(* Logix 5000 project; controller PLC_MCC1300_75F1 vendor 1 type 14 code 166 rev 32.11; software revision 32.04; part 42 of 83 *)
(* tags used below, declared in another part *)
   AUX_xDebugNewPlate : BOOL;
   CM_DATA_Snap_Rx : CM_DATA_Z200;
   CM_INPUT_Z200_Sync : CM_INPUT_Z200;
   CONST_tAux : AUX_COSTANTS;
   CONST_tPlant : UDT_PLANT_CONSTANTS;
   ECL_HLD_AUTO : ALIAS FOR N14[240].2;
   ECL_HLD_AUTO_N : ALIAS FOR I[36].14;
   ECL_HLD_AUTO_S : ALIAS FOR I[80].14;
   ECL_HLD_UP : ALIAS FOR N14[240].3;
   ECL_HLD_UP_N : ALIAS FOR I[36].15;
   ECL_HLD_UP_S : ALIAS FOR I[80].15;
   FL_HLD_AUTO : ALIAS FOR N14[240].0;
   FL_HLD_AUTO_N : ALIAS FOR I[36].12;
   FL_HLD_AUTO_S : ALIAS FOR I[80].12;
   FL_HLD_UP : ALIAS FOR N14[240].1;
   FL_HLD_UP_N : ALIAS FOR I[36].13;
   FL_HLD_UP_S : ALIAS FOR I[80].13;
   GP_OB_InitializeMain : GP_OB_Initialize;
   GP_PlateYPosition : GP_PlateYPosition;
   GP_PosWindow : GP_PosWindow;
   HOLD_DWN_ECLPS : ALIAS FOR O[38].5;
   HOLD_DWN_FLOAT : ALIAS FOR O[38].4;
   I : INT[128];   // Local Input Updates Input Slot 2
   M302SpeedUp : MAC_SpeedUp;
   M302SpeedUp_ALM : MAC_SpeedUp_ALM;
   M302SpeedUp_HMR : MAC_SpeedUp_HMR;
   M302SpeedUp_HMW : MAC_SpeedUp_HMW;
   O : INT[128];
   TMP_dConv : DINT;
   TMP_dConvDebug : DINT;
   TMP_dIndexMotor : DINT;
   TMP_dIndexNext : DINT;
   TMP_dIndexNextDebug : DINT;
   TMP_dIndexPrevious : DINT;
   TMP_dIndexPreviousDebug : DINT;
   TMP_dLehrSpeed : DINT;
   TMP_dLineSpeed : DINT;
   TMP_x : BOOL;
   TMP_xFirstConv : BOOL;
   TMP_xLastConv : BOOL;
   TMP_xLastConvDebug : BOOL;
   xAlwaysOFF : BOOL;
   Z200_SnapDataEth : UDT_ConvoyCap_ZC[2];
   Z300_Conveyor : UDT_StandConv[29];
   Z300_Conveyor_ALM : MAC_Conveyor_ZC_ALM[29];
   Z300_Conveyor_Conf : UDT_Conveyor_Config[29];
   Z300_Conveyor_HMR : MAC_Conveyor_ZC_HMR[29];
   Z300_Conveyor_HMW : MAC_Conveyor_ZC_HMW[29];
   Z300_LineTracking : UDT_LINE_TRACKING;
   Z301 : MAC_Zone_ML;
   Z301_HMR : MAC_Zone_ML_HMR;
   Z301_HMW : MAC_Zone_ML_HMW;
(* MainProgram, continued *)

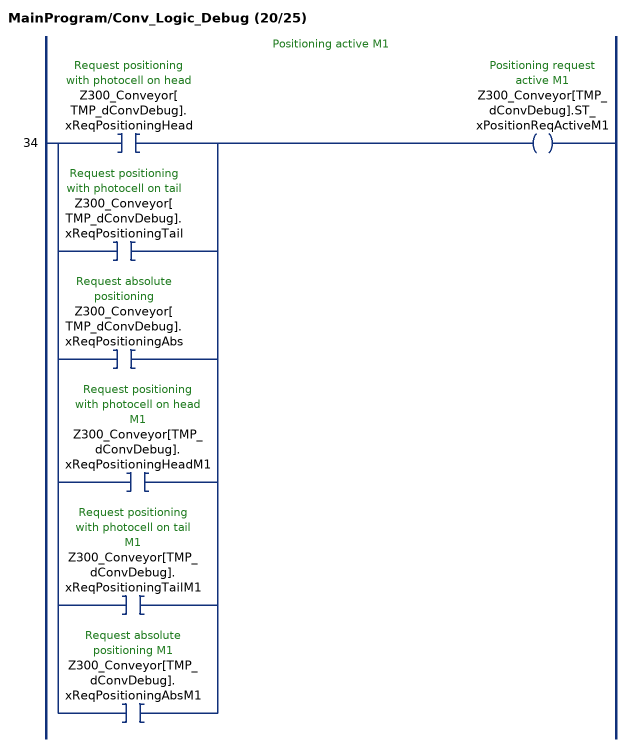
   // Positioning active M1
   34: [XIC(Z300_Conveyor[TMP_dConvDebug].xReqPositioningHead) ,XIC(Z300_Conveyor[TMP_dConvDebug].xReqPositioningTail) ,XIC(Z300_Conveyor[TMP_dConvDebug].xReqPositioningAbs) ,XIC(Z300_Conveyor[TMP_dConvDebug].xReqPositioningHeadM1) ,XIC(Z300_Conveyor[TMP_dConvDebug].xReqPositioningTailM1) ,XIC(Z300_Conveyor[TMP_dConvDebug].xReqPositioningAbsM1) ]OTE(Z300_Conveyor[TMP_dConvDebug].ST_xPositionReqActiveM1);
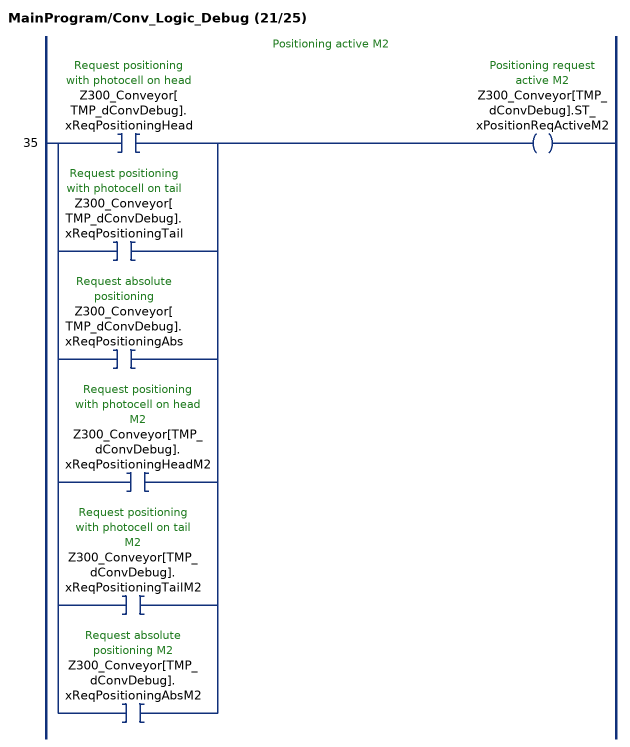
   // Positioning active M2
   35: [XIC(Z300_Conveyor[TMP_dConvDebug].xReqPositioningHead) ,XIC(Z300_Conveyor[TMP_dConvDebug].xReqPositioningTail) ,XIC(Z300_Conveyor[TMP_dConvDebug].xReqPositioningAbs) ,XIC(Z300_Conveyor[TMP_dConvDebug].xReqPositioningHeadM2) ,XIC(Z300_Conveyor[TMP_dConvDebug].xReqPositioningTailM2) ,XIC(Z300_Conveyor[TMP_dConvDebug].xReqPositioningAbsM2) ]OTE(Z300_Conveyor[TMP_dConvDebug].ST_xPositionReqActiveM2);
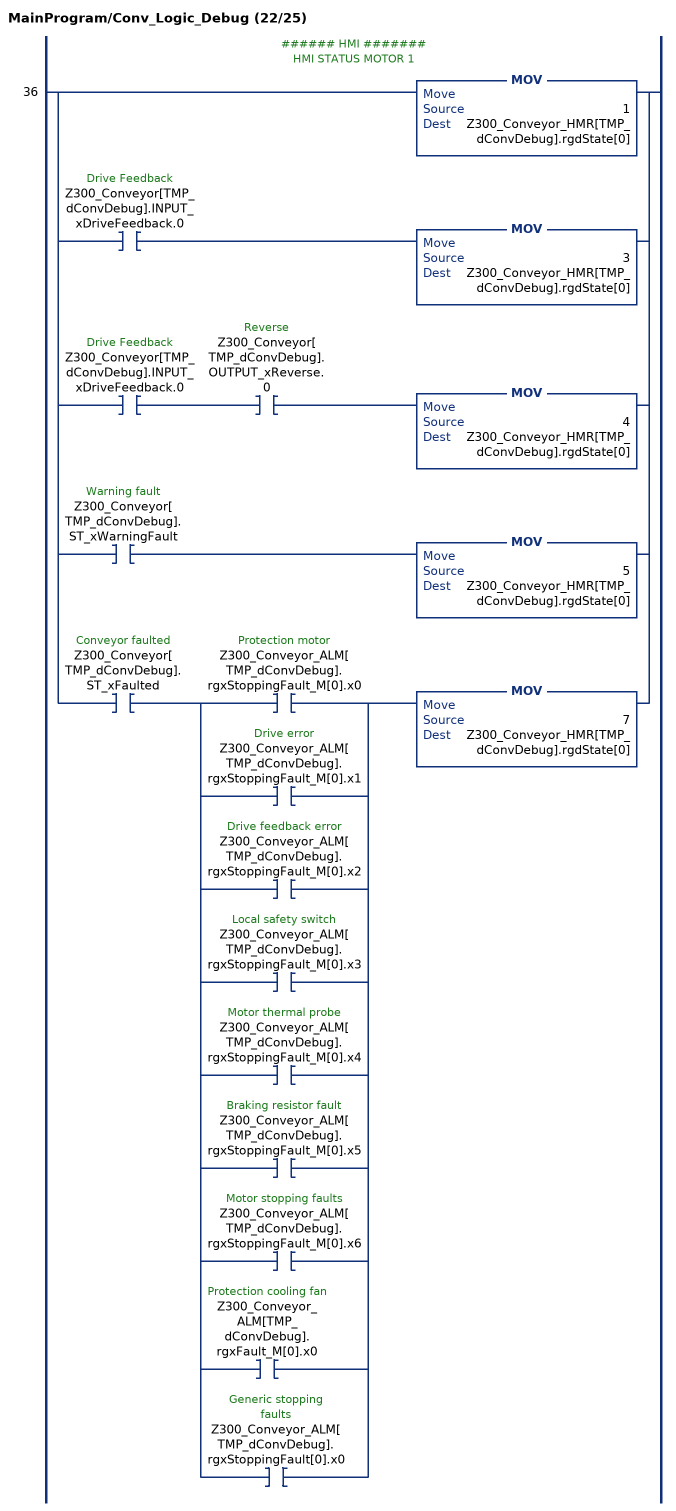
   // ###### HMI #######
   // HMI STATUS MOTOR 1
   36: [MOV(1,Z300_Conveyor_HMR[TMP_dConvDebug].rgdState[0]) ,XIC(Z300_Conveyor[TMP_dConvDebug].INPUT_xDriveFeedback.0) MOV(3,Z300_Conveyor_HMR[TMP_dConvDebug].rgdState[0]) ,XIC(Z300_Conveyor[TMP_dConvDebug].INPUT_xDriveFeedback.0) XIC(Z300_Conveyor[TMP_dConvDebug].OUTPUT_xReverse.0) MOV(4,Z300_Conveyor_HMR[TMP_dConvDebug].rgdState[0]) ,XIC(Z300_Conveyor[TMP_dConvDebug].ST_xWarningFault) MOV(5,Z300_Conveyor_HMR[TMP_dConvDebug].rgdState[0]) ,XIC(Z300_Conveyor[TMP_dConvDebug].ST_xFaulted) [XIC(Z300_Conveyor_ALM[TMP_dConvDebug].rgxStoppingFault_M[0].x0) ,XIC(Z300_Conveyor_ALM[TMP_dConvDebug].rgxStoppingFault_M[0].x1) ,XIC(Z300_Conveyor_ALM[TMP_dConvDebug].rgxStoppingFault_M[0].x2) ,XIC(Z300_Conveyor_ALM[TMP_dConvDebug].rgxStoppingFault_M[0].x3) ,XIC(Z300_Conveyor_ALM[TMP_dConvDebug].rgxStoppingFault_M[0].x4) ,XIC(Z300_Conveyor_ALM[TMP_dConvDebug].rgxStoppingFault_M[0].x5) ,XIC(Z300_Conveyor_ALM[TMP_dConvDebug].rgxStoppingFault_M[0].x6) ,XIC(Z300_Conveyor_ALM[TMP_dConvDebug].rgxFault_M[0].x0) ,XIC(Z300_Conveyor_ALM[TMP_dConvDebug].rgxStoppingFault[0].x0) ] MOV(7,Z300_Conveyor_HMR[TMP_dConvDebug].rgdState[0]) ];
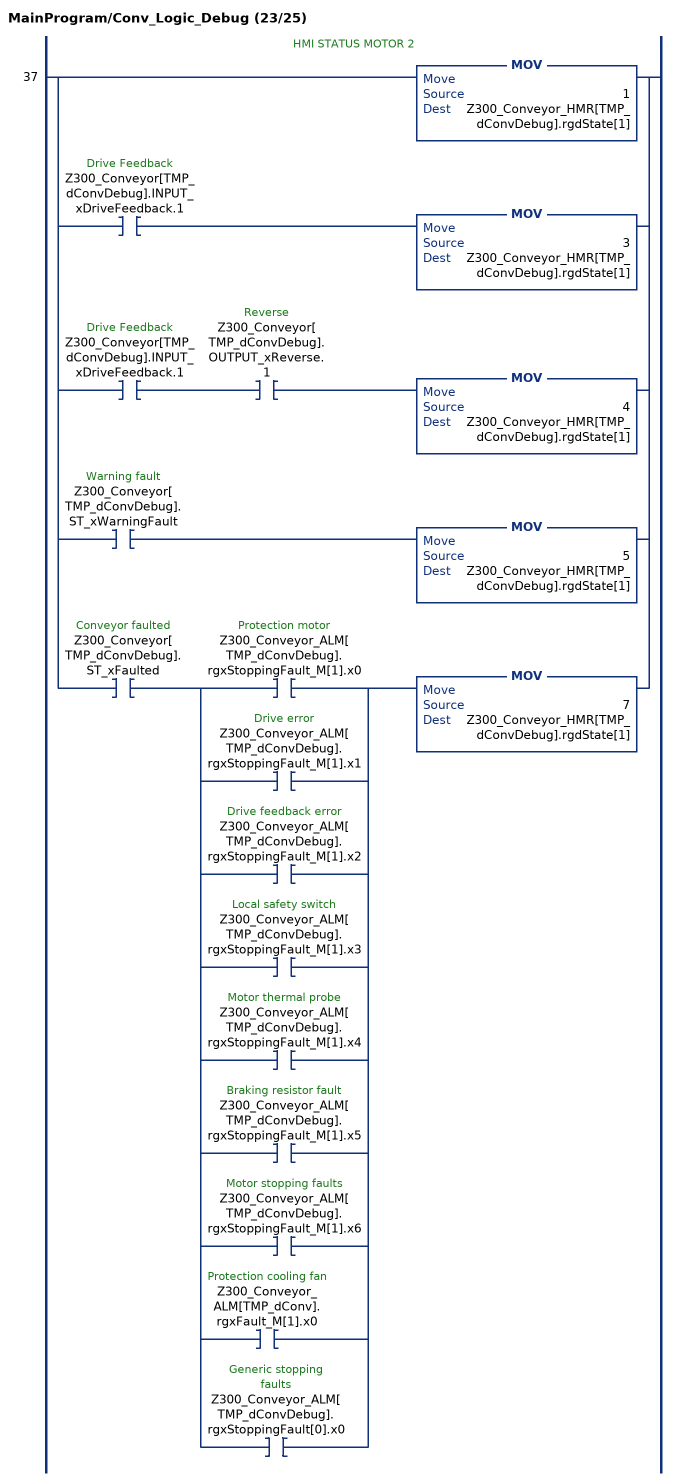
   // HMI STATUS MOTOR 2
   37: [MOV(1,Z300_Conveyor_HMR[TMP_dConvDebug].rgdState[1]) ,XIC(Z300_Conveyor[TMP_dConvDebug].INPUT_xDriveFeedback.1) MOV(3,Z300_Conveyor_HMR[TMP_dConvDebug].rgdState[1]) ,XIC(Z300_Conveyor[TMP_dConvDebug].INPUT_xDriveFeedback.1) XIC(Z300_Conveyor[TMP_dConvDebug].OUTPUT_xReverse.1) MOV(4,Z300_Conveyor_HMR[TMP_dConvDebug].rgdState[1]) ,XIC(Z300_Conveyor[TMP_dConvDebug].ST_xWarningFault) MOV(5,Z300_Conveyor_HMR[TMP_dConvDebug].rgdState[1]) ,XIC(Z300_Conveyor[TMP_dConvDebug].ST_xFaulted) [XIC(Z300_Conveyor_ALM[TMP_dConvDebug].rgxStoppingFault_M[1].x0) ,XIC(Z300_Conveyor_ALM[TMP_dConvDebug].rgxStoppingFault_M[1].x1) ,XIC(Z300_Conveyor_ALM[TMP_dConvDebug].rgxStoppingFault_M[1].x2) ,XIC(Z300_Conveyor_ALM[TMP_dConvDebug].rgxStoppingFault_M[1].x3) ,XIC(Z300_Conveyor_ALM[TMP_dConvDebug].rgxStoppingFault_M[1].x4) ,XIC(Z300_Conveyor_ALM[TMP_dConvDebug].rgxStoppingFault_M[1].x5) ,XIC(Z300_Conveyor_ALM[TMP_dConvDebug].rgxStoppingFault_M[1].x6) ,XIC(Z300_Conveyor_ALM[TMP_dConv].rgxFault_M[1].x0) ,XIC(Z300_Conveyor_ALM[TMP_dConvDebug].rgxStoppingFault[0].x0) ] MOV(7,Z300_Conveyor_HMR[TMP_dConvDebug].rgdState[1]) ];
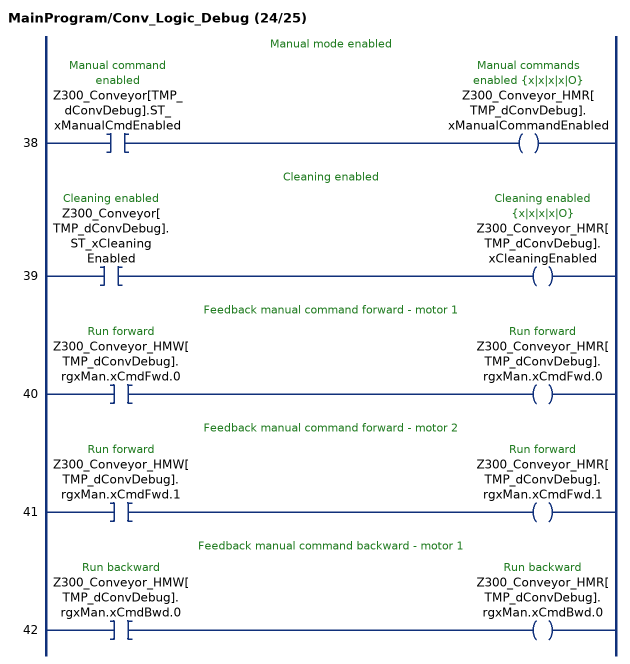
   // Manual mode enabled
   38: XIC(Z300_Conveyor[TMP_dConvDebug].ST_xManualCmdEnabled)OTE(Z300_Conveyor_HMR[TMP_dConvDebug].xManualCommandEnabled);
   // Cleaning enabled
   39: XIC(Z300_Conveyor[TMP_dConvDebug].ST_xCleaningEnabled)OTE(Z300_Conveyor_HMR[TMP_dConvDebug].xCleaningEnabled);
   // Feedback manual command forward - motor 1
   40: XIC(Z300_Conveyor_HMW[TMP_dConvDebug].rgxMan.xCmdFwd.0)OTE(Z300_Conveyor_HMR[TMP_dConvDebug].rgxMan.xCmdFwd.0);
   // Feedback manual command forward - motor 2
   41: XIC(Z300_Conveyor_HMW[TMP_dConvDebug].rgxMan.xCmdFwd.1)OTE(Z300_Conveyor_HMR[TMP_dConvDebug].rgxMan.xCmdFwd.1);
   // Feedback manual command backward - motor 1
   42: XIC(Z300_Conveyor_HMW[TMP_dConvDebug].rgxMan.xCmdBwd.0)OTE(Z300_Conveyor_HMR[TMP_dConvDebug].rgxMan.xCmdBwd.0);
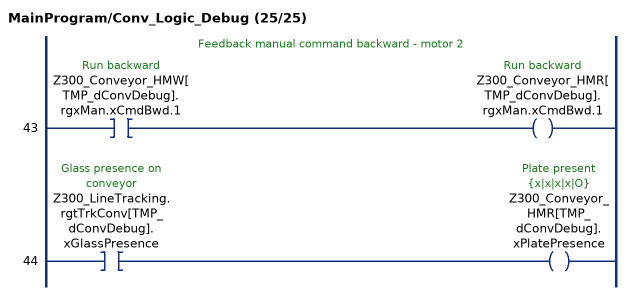
   // Feedback manual command backward - motor 2
   43: XIC(Z300_Conveyor_HMW[TMP_dConvDebug].rgxMan.xCmdBwd.1)OTE(Z300_Conveyor_HMR[TMP_dConvDebug].rgxMan.xCmdBwd.1);
   44: XIC(Z300_LineTracking.rgtTrkConv[TMP_dConvDebug].xGlassPresence)OTE(Z300_Conveyor_HMR[TMP_dConvDebug].xPlatePresence);
END_ROUTINE

ROUTINE Conv_Main   (* structured text *)
   
   //FOR TMP_dConv := 0 TO CONST_tPlant.dNumOfConveyors - 1 DO
   //After the conveyor logic modifications conveyors have to be called from end to begin of the line
   FOR TMP_dConv := CONST_tPlant.dNumOfConveyors - 1 TO 0 BY -1 DO
   
   	JSR(Conv_Faults);
   
   	Z300_Conveyor[TMP_dConv].ST_xOutMotorRun := 1;
   	FOR TMP_dIndexMotor := 0 TO Z300_Conveyor_Conf[TMP_dConv].dMotorNumber DO
   		Z300_Conveyor[TMP_dConv].ST_xOutMotorRun := Z300_Conveyor[TMP_dConv].ST_xOutMotorRun AND Z300_Conveyor[TMP_dConv].OUTPUT_xRun.[TMP_dIndexMotor];
   		Z300_Conveyor[TMP_dConv].ST_rgxOutMotorRunSgm.[TMP_dIndexMotor] := Z300_Conveyor[TMP_dConv].OUTPUT_xRun.[TMP_dIndexMotor];
   	END_FOR;
   
   	//Index Conveyor Previous/Next
   	TMP_xFirstConv := 0;
   	TMP_xLastConv := 0;
   	IF TMP_dConv <=0 THEN
   		TMP_xFirstConv := 1;
   		TMP_dIndexPrevious := TMP_dConv;
   	ELSE
   		TMP_dIndexPrevious := TMP_dConv - 1;
   	END_IF;
   	//Next Conveyor and Last Conveyor
   	//IF TMP_dConv >= CONST_tPlant.dNumOfConveyors - 1 THEN
   	IF TMP_dConv >= CONST_tPlant.dNumOfConveyors - 2 THEN // gli ultimi due convogliatori sono stati uniti
   		TMP_xLastConv := 1;
   		TMP_dIndexNext := TMP_dConv;
   	ELSE
   		TMP_dIndexNext := TMP_dConv + 1;
   	END_IF;
   
   	//Enable control error
   	Z300_Conveyor[TMP_dConv].ST_xEnableControlError := Z300_Conveyor[TMP_dConv].tIN_Zone.xEnableControlError;
   
   	//Feedback, ReadyToMove, Deceleration and position reached of drive
   	Z300_Conveyor[TMP_dConv].ST_xRotationFeedback := 1;
   	Z300_Conveyor[TMP_dConv].ST_xAxleReadyToMoveDelayed := 1;
   	Z300_Conveyor[TMP_dConv].ST_xDriveInDec := 0;
   	Z300_Conveyor[TMP_dConv].ST_xPositionReached := 1;
   	FOR TMP_dIndexMotor := 0 TO Z300_Conveyor_Conf[TMP_dConv].dMotorNumber DO
   		Z300_Conveyor[TMP_dConv].ST_xRotationFeedback := Z300_Conveyor[TMP_dConv].ST_xRotationFeedback AND Z300_Conveyor[TMP_dConv].INPUT_xDriveFeedback.[TMP_dIndexMotor];
   		Z300_Conveyor[TMP_dConv].ST_xAxleReadyToMoveDelayed := Z300_Conveyor[TMP_dConv].ST_xAxleReadyToMoveDelayed AND Z300_Conveyor[TMP_dConv].INPUT_xDriveReady.[TMP_dIndexMotor];
   		Z300_Conveyor[TMP_dConv].ST_xDriveInDec := Z300_Conveyor[TMP_dConv].ST_xDriveInDec AND Z300_Conveyor[TMP_dConv].INPUT_xDriveDeceleration.[TMP_dIndexMotor];
   		Z300_Conveyor[TMP_dConv].ST_xPositionReached := Z300_Conveyor[TMP_dConv].ST_xPositionReached AND Z300_Conveyor[TMP_dConv].INPUT_xDrivePositionReached.[TMP_dIndexMotor];
   
   	END_FOR;
   
   	//Speed value
   	Z300_Conveyor[TMP_dConv].INPUT_rgdRefSpeed_mm_min[0] := Z300_Conveyor[TMP_dConv].tIN_Zone.dAutoSpeed_mm_min;
   	Z300_Conveyor[TMP_dConv].INPUT_rgdRefSpeed_mm_min[1] := Z300_Conveyor[TMP_dConv].tIN_Zone.dLehrSpeed_mm_min;
   	Z300_Conveyor[TMP_dConv].INPUT_rgdRefSpeed_mm_min[2] := Z300_Conveyor[TMP_dConv].tIN_Zone.dCleaningSpeed_mm_min;
   	Z300_Conveyor[TMP_dConv].INPUT_rgdRefSpeed_mm_min[3] := Z300_Conveyor[TMP_dConv].tIN_Zone.dSpecialSpeed_mm_min;
   	Z300_Conveyor[TMP_dConv].INPUT_rgdRefSpeed_mm_min[4] := Z300_Conveyor[TMP_dConv].tIN_Zone.dManualSpeed_mm_min;
   
   	//Acceleration
   	Z300_Conveyor[TMP_dConv].AUX_rgrAcc_m_s2[0] := Z300_Conveyor_Conf[TMP_dConv].rAccH_ms2;
   	Z300_Conveyor[TMP_dConv].AUX_rgrAcc_m_s2[1] := Z300_Conveyor_Conf[TMP_dConv].rAccH_ms2;
   
   	//Deceleration
   	Z300_Conveyor[TMP_dConv].AUX_rgrDec_m_s2[0] := Z300_Conveyor_Conf[TMP_dConv].rDecH_ms2;
   	Z300_Conveyor[TMP_dConv].AUX_rgrDec_m_s2[1] := Z300_Conveyor_Conf[TMP_dConv].rDecH_ms2;
   
   	//Logic
   	IF TMP_dConv = 12 THEN
   		TMP_dConvDebug := TMP_dConv;
   		TMP_dIndexNextDebug := TMP_dIndexNext;
   		TMP_dIndexPreviousDebug := TMP_dIndexPrevious;
   		TMP_xLastConvDebug := TMP_xLastConv;
   		JSR(Conv_Logic_Debug);
   	ELSE
   		JSR(Conv_Logic);
   	END_IF;
   
   END_FOR;
   
END_ROUTINE

ROUTINE Conv_Mapping   (* structured text *)
   
   // Z301
   /*
   FOR TMP_dConv := 0 TO 28 DO
   	Z300_Conveyor[TMP_dConv].tIN_Zone.xCleanZoneAccepted := Z301.ST_xCleaningAccepted;
   	Z300_Conveyor[TMP_dConv].tIN_Zone.xStartCycleRequest := Z301.ST_xStartCycleRequest;
   	Z300_Conveyor[TMP_dConv].tIN_Zone.xCycleON := Z301.ST_xCycleON;
   	Z300_Conveyor[TMP_dConv].tIN_Zone.xManualCmdZoneEnabled := Z301.ST_xManuModeAccepted;
   	Z300_Conveyor[TMP_dConv].tIN_Zone.xResetFault := Z301.ST_xAlarmOff;
   	Z300_Conveyor[TMP_dConv].tIN_Zone.xCmdFwdAll := Z301_HMW.rgxMan.0 OR Z301_HMW.rgxMan.2;
   	Z300_Conveyor[TMP_dConv].tIN_Zone.xCmdBwdAll := Z301_HMW.rgxMan.1 OR Z301_HMW.rgxMan.3;
   	Z300_Conveyor[TMP_dConv].tIN_Zone.dStartCleaning := 0;
   	Z300_Conveyor[TMP_dConv].tIN_Zone.xEnableControlError := Z301.ST_xEnableControlError;
   	Z300_Conveyor[TMP_dConv].tIN_Zone.dAutoSpeed_mm_min := Z301_HMR.dAutoSpeed_mm_min;
   	Z300_Conveyor[TMP_dConv].tIN_Zone.dLehrSpeed_mm_min := Z301.AUX_dLehrSpeed_mm_min;
   	Z300_Conveyor[TMP_dConv].tIN_Zone.dSpecialSpeed_mm_min := Z301_HMR.dAutoSpeedForBreakings_mm_min;
   	Z300_Conveyor[TMP_dConv].tIN_Zone.dManualSpeed_mm_min := Z301_HMR.dManualSpeed_mm_min;
   	Z300_Conveyor[TMP_dConv].tIN_Zone.dCleaningSpeed_mm_min := Z301.AUX_dLehrSpeed_mm_min;
   	Z300_Conveyor[TMP_dConv].tIN_Zone.xExternalConditionCleaning := 1;
   END_FOR;
   */
   //M302-M303
   FOR TMP_dConv := 0 TO 8 DO
   	Z300_Conveyor[TMP_dConv].tIN_Zone.xCleanZoneAccepted := Z301.ST_xCleaningAccepted;
   	Z300_Conveyor[TMP_dConv].tIN_Zone.xStartCycleRequest := Z301.ST_xStartCycleRequest;
   	Z300_Conveyor[TMP_dConv].tIN_Zone.xCycleON := Z301.ST_xCycleON;
   	Z300_Conveyor[TMP_dConv].tIN_Zone.xManualCmdZoneEnabled := Z301.ST_xManuModeAccepted;
   	Z300_Conveyor[TMP_dConv].tIN_Zone.xResetFault := Z301.ST_xAlarmOff;
   	Z300_Conveyor[TMP_dConv].tIN_Zone.xCmdFwdAll := Z301_HMW.rgxMan.0 OR Z301_HMW.rgxMan.2;
   	Z300_Conveyor[TMP_dConv].tIN_Zone.xCmdBwdAll := Z301_HMW.rgxMan.1 OR Z301_HMW.rgxMan.3;
   	Z300_Conveyor[TMP_dConv].tIN_Zone.dStartCleaning := 0;
   	Z300_Conveyor[TMP_dConv].tIN_Zone.xEnableControlError := Z301.ST_xEnableControlError;
   	Z300_Conveyor[TMP_dConv].tIN_Zone.dAutoSpeed_mm_min := Z301.AUX_dLehrSpeed_mm_min;
   	Z300_Conveyor[TMP_dConv].tIN_Zone.dLehrSpeed_mm_min := Z301.AUX_dLehrSpeed_mm_min;
   	Z300_Conveyor[TMP_dConv].tIN_Zone.dSpecialSpeed_mm_min := Z301_HMR.dAutoSpeedForBreakings_mm_min;
   	Z300_Conveyor[TMP_dConv].tIN_Zone.dManualSpeed_mm_min := Z301_HMR.dManualSpeed_mm_min;
   	Z300_Conveyor[TMP_dConv].tIN_Zone.dCleaningSpeed_mm_min := Z301.AUX_dLehrSpeed_mm_min;
   	Z300_Conveyor[TMP_dConv].tIN_Zone.xExternalConditionCleaning := 1;
   END_FOR;
   
   //M304-M305-M306
   FOR TMP_dConv := 9 TO 11 DO
   	Z300_Conveyor[TMP_dConv].tIN_Zone.xCleanZoneAccepted := Z301.ST_xCleaningAccepted;
   	Z300_Conveyor[TMP_dConv].tIN_Zone.xStartCycleRequest := Z301.ST_xStartCycleRequest;
   	Z300_Conveyor[TMP_dConv].tIN_Zone.xCycleON := Z301.ST_xCycleON;
   	Z300_Conveyor[TMP_dConv].tIN_Zone.xManualCmdZoneEnabled := Z301.ST_xManuModeAccepted;
   	Z300_Conveyor[TMP_dConv].tIN_Zone.xResetFault := Z301.ST_xAlarmOff;
   	Z300_Conveyor[TMP_dConv].tIN_Zone.xCmdFwdAll := Z301_HMW.rgxMan.0 OR Z301_HMW.rgxMan.2;
   	Z300_Conveyor[TMP_dConv].tIN_Zone.xCmdBwdAll := Z301_HMW.rgxMan.1 OR Z301_HMW.rgxMan.3;
   	Z300_Conveyor[TMP_dConv].tIN_Zone.dStartCleaning := 0;
   	Z300_Conveyor[TMP_dConv].tIN_Zone.xEnableControlError := Z301.ST_xEnableControlError;
   	Z300_Conveyor[TMP_dConv].tIN_Zone.dAutoSpeed_mm_min :=Z301_HMR.dAutoSpeedForBreakings_mm_min;
   	Z300_Conveyor[TMP_dConv].tIN_Zone.dLehrSpeed_mm_min := Z301.AUX_dLehrSpeed_mm_min;
   	Z300_Conveyor[TMP_dConv].tIN_Zone.dSpecialSpeed_mm_min := Z301_HMR.dAutoSpeedForBreakings_mm_min;
   	Z300_Conveyor[TMP_dConv].tIN_Zone.dManualSpeed_mm_min := Z301_HMR.dManualSpeed_mm_min;
   	Z300_Conveyor[TMP_dConv].tIN_Zone.dCleaningSpeed_mm_min := Z301.AUX_dLehrSpeed_mm_min;
   	Z300_Conveyor[TMP_dConv].tIN_Zone.xExternalConditionCleaning := 1;
   END_FOR;
   
   //M307A-B-C
   FOR TMP_dConv := 12 TO 17 DO
   	Z300_Conveyor[TMP_dConv].tIN_Zone.xCleanZoneAccepted := Z301.ST_xCleaningAccepted;
   	Z300_Conveyor[TMP_dConv].tIN_Zone.xStartCycleRequest := Z301.ST_xStartCycleRequest;
   	Z300_Conveyor[TMP_dConv].tIN_Zone.xCycleON := Z301.ST_xCycleON;
   	Z300_Conveyor[TMP_dConv].tIN_Zone.xManualCmdZoneEnabled := Z301.ST_xManuModeAccepted;
   	Z300_Conveyor[TMP_dConv].tIN_Zone.xResetFault := Z301.ST_xAlarmOff;
   	Z300_Conveyor[TMP_dConv].tIN_Zone.xCmdFwdAll := Z301_HMW.rgxMan.0 OR Z301_HMW.rgxMan.2;
   	Z300_Conveyor[TMP_dConv].tIN_Zone.xCmdBwdAll := Z301_HMW.rgxMan.1 OR Z301_HMW.rgxMan.3;
   	Z300_Conveyor[TMP_dConv].tIN_Zone.dStartCleaning := 0;
   	Z300_Conveyor[TMP_dConv].tIN_Zone.xEnableControlError := Z301.ST_xEnableControlError;
   	Z300_Conveyor[TMP_dConv].tIN_Zone.dAutoSpeed_mm_min :=Z301_HMR.dAutoSpeedForBreakings_mm_min;
   	Z300_Conveyor[TMP_dConv].tIN_Zone.dLehrSpeed_mm_min := Z301_HMR.dAutoSpeedForBreakings_mm_min;
   	Z300_Conveyor[TMP_dConv].tIN_Zone.dSpecialSpeed_mm_min := Z301_HMR.dAutoSpeed_mm_min;
   	Z300_Conveyor[TMP_dConv].tIN_Zone.dManualSpeed_mm_min := Z301_HMR.dManualSpeed_mm_min;
   	Z300_Conveyor[TMP_dConv].tIN_Zone.dCleaningSpeed_mm_min := Z301.AUX_dLehrSpeed_mm_min;
   	Z300_Conveyor[TMP_dConv].tIN_Zone.xExternalConditionCleaning := 1;
   END_FOR;
   
   //FROM M307D TO M315M3
   FOR TMP_dConv := 18 TO 28 DO
   	Z300_Conveyor[TMP_dConv].tIN_Zone.xCleanZoneAccepted := Z301.ST_xCleaningAccepted;
   	Z300_Conveyor[TMP_dConv].tIN_Zone.xStartCycleRequest := Z301.ST_xStartCycleRequest;
   	Z300_Conveyor[TMP_dConv].tIN_Zone.xCycleON := Z301.ST_xCycleON;
   	Z300_Conveyor[TMP_dConv].tIN_Zone.xManualCmdZoneEnabled := Z301.ST_xManuModeAccepted;
   	Z300_Conveyor[TMP_dConv].tIN_Zone.xResetFault := Z301.ST_xAlarmOff;
   	Z300_Conveyor[TMP_dConv].tIN_Zone.xCmdFwdAll := Z301_HMW.rgxMan.0 OR Z301_HMW.rgxMan.2;
   	Z300_Conveyor[TMP_dConv].tIN_Zone.xCmdBwdAll := Z301_HMW.rgxMan.1 OR Z301_HMW.rgxMan.3;
   	Z300_Conveyor[TMP_dConv].tIN_Zone.dStartCleaning := 0;
   	Z300_Conveyor[TMP_dConv].tIN_Zone.xEnableControlError := Z301.ST_xEnableControlError;
   	Z300_Conveyor[TMP_dConv].tIN_Zone.dAutoSpeed_mm_min := Z301_HMR.dAutoSpeed_mm_min;
   	Z300_Conveyor[TMP_dConv].tIN_Zone.dLehrSpeed_mm_min := Z301.AUX_dLehrSpeed_mm_min;
   	Z300_Conveyor[TMP_dConv].tIN_Zone.dSpecialSpeed_mm_min := Z301_HMR.dAutoSpeed_mm_min;
   	Z300_Conveyor[TMP_dConv].tIN_Zone.dManualSpeed_mm_min := Z301_HMR.dManualSpeed_mm_min;
   	Z300_Conveyor[TMP_dConv].tIN_Zone.dCleaningSpeed_mm_min := Z301.AUX_dLehrSpeed_mm_min;
   	Z300_Conveyor[TMP_dConv].tIN_Zone.xExternalConditionCleaning := 1;
   END_FOR;
   
   
   
   //If M323 popup not low cannot clean M323
   //Z300_Conveyor[21].tIN_Zone.xExternalConditionCleaning := M323Popup.INPUT_xPopupLow;
   //If M327 popup not low cannot clean M327
   //Z300_Conveyor[26].tIN_Zone.xExternalConditionCleaning := M327Popup.INPUT_xPopupLow;
   
END_ROUTINE

ROUTINE Hold_Down_Wheels   (* ladder *)
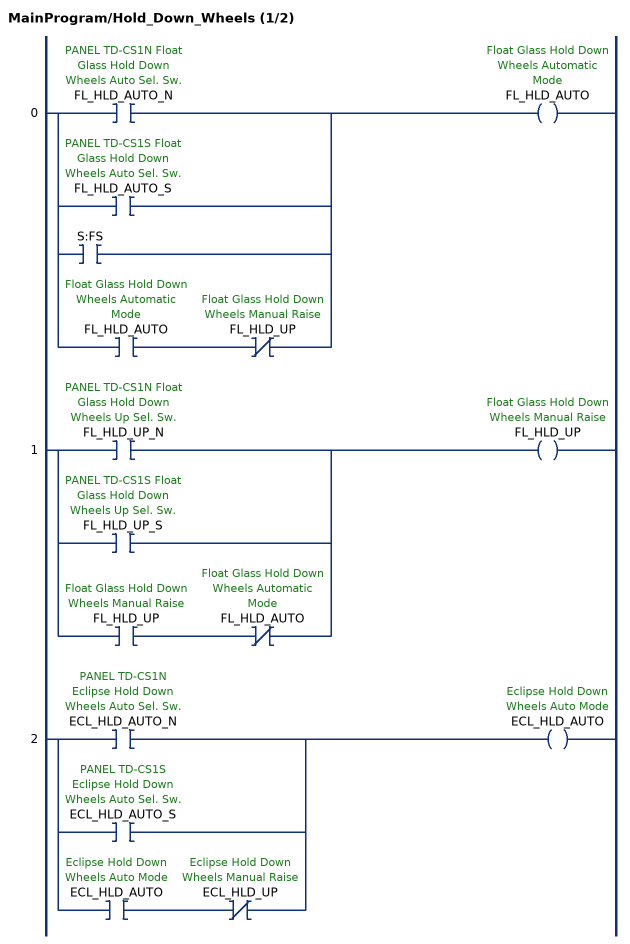
   0: [[XIC(FL_HLD_AUTO_N) ,XIC(FL_HLD_AUTO_S) ,XIC(S:FS) ] ,XIC(FL_HLD_AUTO) XIO(FL_HLD_UP) ]OTE(FL_HLD_AUTO);
   1: [[XIC(FL_HLD_UP_N) ,XIC(FL_HLD_UP_S) ] ,XIC(FL_HLD_UP) XIO(FL_HLD_AUTO) ]OTE(FL_HLD_UP);
   2: [[XIC(ECL_HLD_AUTO_N) ,XIC(ECL_HLD_AUTO_S) ] ,XIC(ECL_HLD_AUTO) XIO(ECL_HLD_UP) ]OTE(ECL_HLD_AUTO);
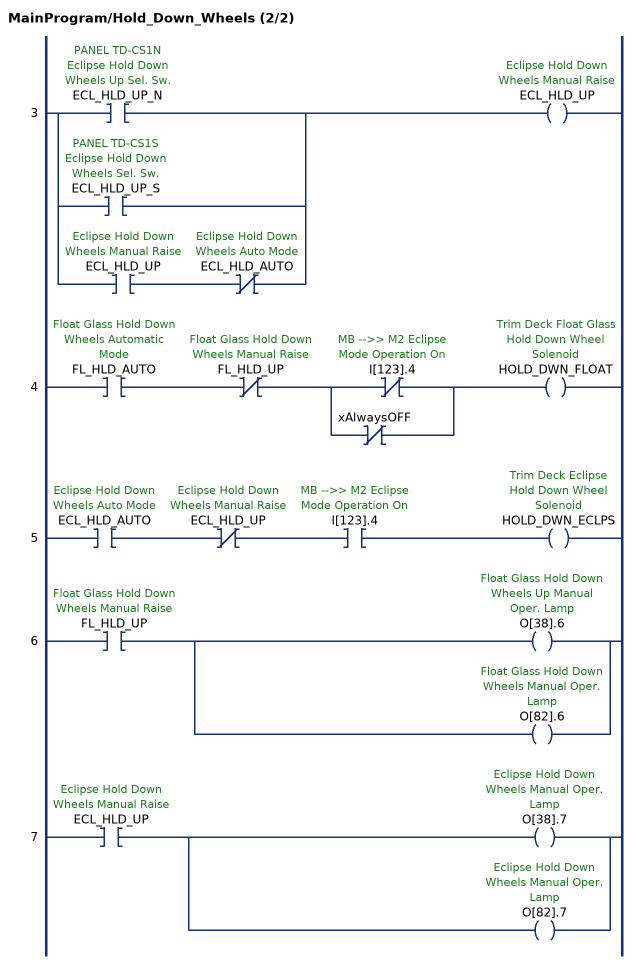
   3: [[XIC(ECL_HLD_UP_N) ,XIC(ECL_HLD_UP_S) ] ,XIC(ECL_HLD_UP) XIO(ECL_HLD_AUTO) ]OTE(ECL_HLD_UP);
   4: XIC(FL_HLD_AUTO)XIO(FL_HLD_UP)[XIO(I[123].4) ,XIO(xAlwaysOFF) ]OTE(HOLD_DWN_FLOAT);
   5: XIC(ECL_HLD_AUTO)XIO(ECL_HLD_UP)XIC(I[123].4)OTE(HOLD_DWN_ECLPS);
   6: XIC(FL_HLD_UP)[OTE(O[38].6) ,OTE(O[82].6) ];
   7: XIC(ECL_HLD_UP)[OTE(O[38].7) ,OTE(O[82].7) ];
END_ROUTINE

ROUTINE inputs_update   (* ladder *)
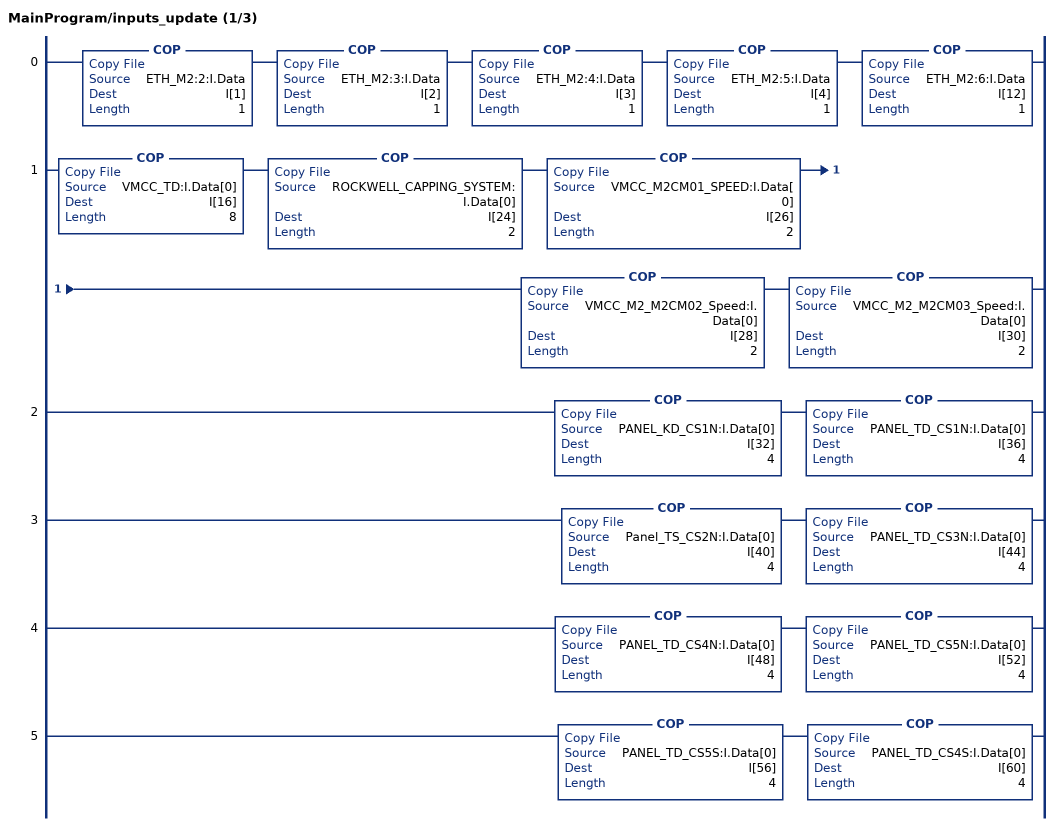
   0: COP(ETH_M2:2:I.Data,I[1],1)COP(ETH_M2:3:I.Data,I[2],1)COP(ETH_M2:4:I.Data,I[3],1)COP(ETH_M2:5:I.Data,I[4],1)COP(ETH_M2:6:I.Data,I[12],1);
   1: COP(VMCC_TD:I.Data[0],I[16],8)COP(ROCKWELL_CAPPING_SYSTEM:I.Data[0],I[24],2)COP(VMCC_M2CM01_SPEED:I.Data[0],I[26],2)COP(VMCC_M2_M2CM02_Speed:I.Data[0],I[28],2)COP(VMCC_M2_M2CM03_Speed:I.Data[0],I[30],2);
   2: COP(PANEL_KD_CS1N:I.Data[0],I[32],4)COP(PANEL_TD_CS1N:I.Data[0],I[36],4);
   3: COP(Panel_TS_CS2N:I.Data[0],I[40],4)COP(PANEL_TD_CS3N:I.Data[0],I[44],4);
   4: COP(PANEL_TD_CS4N:I.Data[0],I[48],4)COP(PANEL_TD_CS5N:I.Data[0],I[52],4);
   5: COP(PANEL_TD_CS5S:I.Data[0],I[56],4)COP(PANEL_TD_CS4S:I.Data[0],I[60],4);